(* Logix 5000 project; controller POA Emulate 5570 rev 30.12; software revision 30.00; part 4 of 6 *)
(* tags used below, declared in another part *)
   Chaskey_Message : DINT[256];
   Chaskey_mlen : DINT;
   Chaskey_MsgBitLen : DINT;
   Chaskey_round : DINT;
   Chaskey_tag : DINT[4];
   Date_time : DINT[7];
   OWF_Add_c : DINT;
   OWF_i : DINT;
   OWF_Input : DINT[17];
   OWF_InputLen : DINT;
   OWF_InputMaxInd : DINT;
   OWF_Result : DINT[17];
   POA_Chain_NM : DINT;
   POA_CKP : DINT[17];
   POA_i : DINT;
   POA_Ins_NM : DINT;
   POA_j : DINT;
   POA_k : DINT;
   POA_lr : DINT;
   POA_m : DINT;
   POA_Microsecond1 : DINT;
   POA_Microsecond2 : DINT;
   POA_MicrosecondABS : DINT;
   POA_OTS : SINT[256,256];
   POA_Pf : DINT[17];
   POA_Pf_Indx : DINT;
   POA_SC_Interval : DINT;
   POA_Second1 : DINT;
   POA_Second2 : DINT;
   POA_SecondABS : DINT;
   POA_SIG_i : DINT;
   POA_tag : DINT[4];
   POA_Vrf_Points : DINT[260,17];
   PRG_Counter : DINT[2];
   PRG_i : DINT;
   PRG_j : DINT;
   PRG_Res_Len : DINT;
   PRG_Result : DINT[128];
   SCAN_CYCLE_TIME : DINT;
   UOWHF_Add_c : DINT;
   UOWHF_Msg : DINT[17];
   UOWHF_Result : DINT[17];
   UOWHF_Vary_Message : DINT[3000];
   UOWHF_Vary_MsgLen : DINT;
   UOWHF_Ver : DINT;
(* MainProgram, continued *)

   		OWF_Add_c.1:=OWF_Result[1].31;
   		OWF_Result[1].31:=0;
   		OWF_Result[2]:=OWF_Result[2] + 102357735+OWF_Add_c;
   		OWF_Add_c.2:=OWF_Result[2].31;
   		OWF_Result[2].31:=0;
   		OWF_Result[3]:=OWF_Result[3] + 1548947751+OWF_Add_c;
   		OWF_Add_c.3:=OWF_Result[3].31;
   		OWF_Result[3].31:=0;
   		OWF_Result[4]:=OWF_Result[4] + 1541273950+OWF_Add_c;
   		OWF_Add_c.4:=OWF_Result[4].31;
   		OWF_Result[4].31:=0;
   		OWF_Result[5]:=OWF_Result[5] + 1965581916+OWF_Add_c;
   		OWF_Add_c.5:=OWF_Result[5].31;
   		OWF_Result[5].31:=0;
   		OWF_Result[6]:=OWF_Result[6] + 714783171+OWF_Add_c;
   		OWF_Add_c.6:=OWF_Result[6].31;
   		OWF_Result[6].31:=0;
   		OWF_Result[7]:=OWF_Result[7] + 952638591+OWF_Add_c;
   		OWF_Add_c.7:=OWF_Result[7].31;
   		OWF_Result[7].31:=0;
   		OWF_Result[8]:=OWF_Result[8] + 1892750752+OWF_Add_c;
   		OWF_Add_c.8:=OWF_Result[8].31;
   		OWF_Result[8].31:=0;
   	End_If;
   	If OWF_Input[7].[20] Then
   		OWF_Result[0]:=OWF_Result[0] + 1923601846+OWF_Add_c;
   		OWF_Add_c.0:=OWF_Result[0].31;
   		OWF_Result[0].31:=0;
   		OWF_Result[1]:=OWF_Result[1] + 431367542+OWF_Add_c;
   		OWF_Add_c.1:=OWF_Result[1].31;
   		OWF_Result[1].31:=0;
   		OWF_Result[2]:=OWF_Result[2] + 812772690+OWF_Add_c;
   		OWF_Add_c.2:=OWF_Result[2].31;
   		OWF_Result[2].31:=0;
   		OWF_Result[3]:=OWF_Result[3] + 1612004830+OWF_Add_c;
   		OWF_Add_c.3:=OWF_Result[3].31;
   		OWF_Result[3].31:=0;
   		OWF_Result[4]:=OWF_Result[4] + 1503607425+OWF_Add_c;
   		OWF_Add_c.4:=OWF_Result[4].31;
   		OWF_Result[4].31:=0;
   		OWF_Result[5]:=OWF_Result[5] + 257117095+OWF_Add_c;
   		OWF_Add_c.5:=OWF_Result[5].31;
   		OWF_Result[5].31:=0;
   		OWF_Result[6]:=OWF_Result[6] + 1165565758+OWF_Add_c;
   		OWF_Add_c.6:=OWF_Result[6].31;
   		OWF_Result[6].31:=0;
   		OWF_Result[7]:=OWF_Result[7] + 1791078952+OWF_Add_c;
   		OWF_Add_c.7:=OWF_Result[7].31;
   		OWF_Result[7].31:=0;
   		OWF_Result[8]:=OWF_Result[8] + 1316586480+OWF_Add_c;
   		OWF_Add_c.8:=OWF_Result[8].31;
   		OWF_Result[8].31:=0;
   	End_If;
   	If OWF_Input[7].[21] Then
   		OWF_Result[0]:=OWF_Result[0] + 1179130031+OWF_Add_c;
   		OWF_Add_c.0:=OWF_Result[0].31;
   		OWF_Result[0].31:=0;
   		OWF_Result[1]:=OWF_Result[1] + 1413483742+OWF_Add_c;
   		OWF_Add_c.1:=OWF_Result[1].31;
   		OWF_Result[1].31:=0;
   		OWF_Result[2]:=OWF_Result[2] + 2076538493+OWF_Add_c;
   		OWF_Add_c.2:=OWF_Result[2].31;
   		OWF_Result[2].31:=0;
   		OWF_Result[3]:=OWF_Result[3] + 415974763+OWF_Add_c;
   		OWF_Add_c.3:=OWF_Result[3].31;
   		OWF_Result[3].31:=0;
   		OWF_Result[4]:=OWF_Result[4] + 461079233+OWF_Add_c;
   		OWF_Add_c.4:=OWF_Result[4].31;
   		OWF_Result[4].31:=0;
   		OWF_Result[5]:=OWF_Result[5] + 207770264+OWF_Add_c;
   		OWF_Add_c.5:=OWF_Result[5].31;
   		OWF_Result[5].31:=0;
   		OWF_Result[6]:=OWF_Result[6] + 670532004+OWF_Add_c;
   		OWF_Add_c.6:=OWF_Result[6].31;
   		OWF_Result[6].31:=0;
   		OWF_Result[7]:=OWF_Result[7] + 164283060+OWF_Add_c;
   		OWF_Add_c.7:=OWF_Result[7].31;
   		OWF_Result[7].31:=0;
   		OWF_Result[8]:=OWF_Result[8] + 1512816438+OWF_Add_c;
   		OWF_Add_c.8:=OWF_Result[8].31;
   		OWF_Result[8].31:=0;
   	End_If;
   	If OWF_Input[7].[22] Then
   		OWF_Result[0]:=OWF_Result[0] + 1897360171+OWF_Add_c;
   		OWF_Add_c.0:=OWF_Result[0].31;
   		OWF_Result[0].31:=0;
   		OWF_Result[1]:=OWF_Result[1] + 1308779824+OWF_Add_c;
   		OWF_Add_c.1:=OWF_Result[1].31;
   		OWF_Result[1].31:=0;
   		OWF_Result[2]:=OWF_Result[2] + 1875593423+OWF_Add_c;
   		OWF_Add_c.2:=OWF_Result[2].31;
   		OWF_Result[2].31:=0;
   		OWF_Result[3]:=OWF_Result[3] + 571271217+OWF_Add_c;
   		OWF_Add_c.3:=OWF_Result[3].31;
   		OWF_Result[3].31:=0;
   		OWF_Result[4]:=OWF_Result[4] + 344940971+OWF_Add_c;
   		OWF_Add_c.4:=OWF_Result[4].31;
   		OWF_Result[4].31:=0;
   		OWF_Result[5]:=OWF_Result[5] + 75339231+OWF_Add_c;
   		OWF_Add_c.5:=OWF_Result[5].31;
   		OWF_Result[5].31:=0;
   		OWF_Result[6]:=OWF_Result[6] + 1428316860+OWF_Add_c;
   		OWF_Add_c.6:=OWF_Result[6].31;
   		OWF_Result[6].31:=0;
   		OWF_Result[7]:=OWF_Result[7] + 1811603075+OWF_Add_c;
   		OWF_Add_c.7:=OWF_Result[7].31;
   		OWF_Result[7].31:=0;
   		OWF_Result[8]:=OWF_Result[8] + 1679786029+OWF_Add_c;
   		OWF_Add_c.8:=OWF_Result[8].31;
   		OWF_Result[8].31:=0;
   	End_If;
   	If OWF_Input[7].[23] Then
   		OWF_Result[0]:=OWF_Result[0] + 271831917+OWF_Add_c;
   		OWF_Add_c.0:=OWF_Result[0].31;
   		OWF_Result[0].31:=0;
   		OWF_Result[1]:=OWF_Result[1] + 663117307+OWF_Add_c;
   		OWF_Add_c.1:=OWF_Result[1].31;
   		OWF_Result[1].31:=0;
   		OWF_Result[2]:=OWF_Result[2] + 1802435718+OWF_Add_c;
   		OWF_Add_c.2:=OWF_Result[2].31;
   		OWF_Result[2].31:=0;
   		OWF_Result[3]:=OWF_Result[3] + 585874673+OWF_Add_c;
   		OWF_Add_c.3:=OWF_Result[3].31;
   		OWF_Result[3].31:=0;
   		OWF_Result[4]:=OWF_Result[4] + 701698092+OWF_Add_c;
   		OWF_Add_c.4:=OWF_Result[4].31;
   		OWF_Result[4].31:=0;
   		OWF_Result[5]:=OWF_Result[5] + 1402770880+OWF_Add_c;
   		OWF_Add_c.5:=OWF_Result[5].31;
   		OWF_Result[5].31:=0;
   		OWF_Result[6]:=OWF_Result[6] + 452824658+OWF_Add_c;
   		OWF_Add_c.6:=OWF_Result[6].31;
   		OWF_Result[6].31:=0;
   		OWF_Result[7]:=OWF_Result[7] + 1400742763+OWF_Add_c;
   		OWF_Add_c.7:=OWF_Result[7].31;
   		OWF_Result[7].31:=0;
   		OWF_Result[8]:=OWF_Result[8] + 2073024045+OWF_Add_c;
   		OWF_Add_c.8:=OWF_Result[8].31;
   		OWF_Result[8].31:=0;
   	End_If;
   	If OWF_Input[7].[24] Then
   		OWF_Result[0]:=OWF_Result[0] + 1367845667+OWF_Add_c;
   		OWF_Add_c.0:=OWF_Result[0].31;
   		OWF_Result[0].31:=0;
   		OWF_Result[1]:=OWF_Result[1] + 1195094582+OWF_Add_c;
   		OWF_Add_c.1:=OWF_Result[1].31;
   		OWF_Result[1].31:=0;
   		OWF_Result[2]:=OWF_Result[2] + 494736933+OWF_Add_c;
   		OWF_Add_c.2:=OWF_Result[2].31;
   		OWF_Result[2].31:=0;
   		OWF_Result[3]:=OWF_Result[3] + 1875737261+OWF_Add_c;
   		OWF_Add_c.3:=OWF_Result[3].31;
   		OWF_Result[3].31:=0;
   		OWF_Result[4]:=OWF_Result[4] + 726339725+OWF_Add_c;
   		OWF_Add_c.4:=OWF_Result[4].31;
   		OWF_Result[4].31:=0;
   		OWF_Result[5]:=OWF_Result[5] + 1862851936+OWF_Add_c;
   		OWF_Add_c.5:=OWF_Result[5].31;
   		OWF_Result[5].31:=0;
   		OWF_Result[6]:=OWF_Result[6] + 296798862+OWF_Add_c;
   		OWF_Add_c.6:=OWF_Result[6].31;
   		OWF_Result[6].31:=0;
   		OWF_Result[7]:=OWF_Result[7] + 1485306441+OWF_Add_c;
   		OWF_Add_c.7:=OWF_Result[7].31;
   		OWF_Result[7].31:=0;
   		OWF_Result[8]:=OWF_Result[8] + 79244469+OWF_Add_c;
   		OWF_Add_c.8:=OWF_Result[8].31;
   		OWF_Result[8].31:=0;
   	End_If;
   	If OWF_Input[7].[25] Then
   		OWF_Result[0]:=OWF_Result[0] + 1748009068+OWF_Add_c;
   		OWF_Add_c.0:=OWF_Result[0].31;
   		OWF_Result[0].31:=0;
   		OWF_Result[1]:=OWF_Result[1] + 153673379+OWF_Add_c;
   		OWF_Add_c.1:=OWF_Result[1].31;
   		OWF_Result[1].31:=0;
   		OWF_Result[2]:=OWF_Result[2] + 1563899973+OWF_Add_c;
   		OWF_Add_c.2:=OWF_Result[2].31;
   		OWF_Result[2].31:=0;
   		OWF_Result[3]:=OWF_Result[3] + 210477071+OWF_Add_c;
   		OWF_Add_c.3:=OWF_Result[3].31;
   		OWF_Result[3].31:=0;
   		OWF_Result[4]:=OWF_Result[4] + 598591903+OWF_Add_c;
   		OWF_Add_c.4:=OWF_Result[4].31;
   		OWF_Result[4].31:=0;
   		OWF_Result[5]:=OWF_Result[5] + 889903791+OWF_Add_c;
   		OWF_Add_c.5:=OWF_Result[5].31;
   		OWF_Result[5].31:=0;
   		OWF_Result[6]:=OWF_Result[6] + 1087681228+OWF_Add_c;
   		OWF_Add_c.6:=OWF_Result[6].31;
   		OWF_Result[6].31:=0;
   		OWF_Result[7]:=OWF_Result[7] + 146945819+OWF_Add_c;
   		OWF_Add_c.7:=OWF_Result[7].31;
   		OWF_Result[7].31:=0;
   		OWF_Result[8]:=OWF_Result[8] + 658778953+OWF_Add_c;
   		OWF_Add_c.8:=OWF_Result[8].31;
   		OWF_Result[8].31:=0;
   	End_If;
   	If OWF_Input[7].[26] Then
   		OWF_Result[0]:=OWF_Result[0] + 1388889236+OWF_Add_c;
   		OWF_Add_c.0:=OWF_Result[0].31;
   		OWF_Result[0].31:=0;
   		OWF_Result[1]:=OWF_Result[1] + 1854230592+OWF_Add_c;
   		OWF_Add_c.1:=OWF_Result[1].31;
   		OWF_Result[1].31:=0;
   		OWF_Result[2]:=OWF_Result[2] + 1952659775+OWF_Add_c;
   		OWF_Add_c.2:=OWF_Result[2].31;
   		OWF_Result[2].31:=0;
   		OWF_Result[3]:=OWF_Result[3] + 693016622+OWF_Add_c;
   		OWF_Add_c.3:=OWF_Result[3].31;
   		OWF_Result[3].31:=0;
   		OWF_Result[4]:=OWF_Result[4] + 19961190+OWF_Add_c;
   		OWF_Add_c.4:=OWF_Result[4].31;
   		OWF_Result[4].31:=0;
   		OWF_Result[5]:=OWF_Result[5] + 1155238848+OWF_Add_c;
   		OWF_Add_c.5:=OWF_Result[5].31;
   		OWF_Result[5].31:=0;
   		OWF_Result[6]:=OWF_Result[6] + 1721973623+OWF_Add_c;
   		OWF_Add_c.6:=OWF_Result[6].31;
   		OWF_Result[6].31:=0;
   		OWF_Result[7]:=OWF_Result[7] + 1298626904+OWF_Add_c;
   		OWF_Add_c.7:=OWF_Result[7].31;
   		OWF_Result[7].31:=0;
   		OWF_Result[8]:=OWF_Result[8] + 704184103+OWF_Add_c;
   		OWF_Add_c.8:=OWF_Result[8].31;
   		OWF_Result[8].31:=0;
   	End_If;
   	If OWF_Input[7].[27] Then
   		OWF_Result[0]:=OWF_Result[0] + 1064559134+OWF_Add_c;
   		OWF_Add_c.0:=OWF_Result[0].31;
   		OWF_Result[0].31:=0;
   		OWF_Result[1]:=OWF_Result[1] + 628496468+OWF_Add_c;
   		OWF_Add_c.1:=OWF_Result[1].31;
   		OWF_Result[1].31:=0;
   		OWF_Result[2]:=OWF_Result[2] + 1741787667+OWF_Add_c;
   		OWF_Add_c.2:=OWF_Result[2].31;
   		OWF_Result[2].31:=0;
   		OWF_Result[3]:=OWF_Result[3] + 650880797+OWF_Add_c;
   		OWF_Add_c.3:=OWF_Result[3].31;
   		OWF_Result[3].31:=0;
   		OWF_Result[4]:=OWF_Result[4] + 927193641+OWF_Add_c;
   		OWF_Add_c.4:=OWF_Result[4].31;
   		OWF_Result[4].31:=0;
   		OWF_Result[5]:=OWF_Result[5] + 690779087+OWF_Add_c;
   		OWF_Add_c.5:=OWF_Result[5].31;
   		OWF_Result[5].31:=0;
   		OWF_Result[6]:=OWF_Result[6] + 1387171811+OWF_Add_c;
   		OWF_Add_c.6:=OWF_Result[6].31;
   		OWF_Result[6].31:=0;
   		OWF_Result[7]:=OWF_Result[7] + 1642242275+OWF_Add_c;
   		OWF_Add_c.7:=OWF_Result[7].31;
   		OWF_Result[7].31:=0;
   		OWF_Result[8]:=OWF_Result[8] + 750154437+OWF_Add_c;
   		OWF_Add_c.8:=OWF_Result[8].31;
   		OWF_Result[8].31:=0;
   	End_If;
   	If OWF_Input[7].[28] Then
   		OWF_Result[0]:=OWF_Result[0] + 1648370074+OWF_Add_c;
   		OWF_Add_c.0:=OWF_Result[0].31;
   		OWF_Result[0].31:=0;
   		OWF_Result[1]:=OWF_Result[1] + 242619355+OWF_Add_c;
   		OWF_Add_c.1:=OWF_Result[1].31;
   		OWF_Result[1].31:=0;
   		OWF_Result[2]:=OWF_Result[2] + 1874736599+OWF_Add_c;
   		OWF_Add_c.2:=OWF_Result[2].31;
   		OWF_Result[2].31:=0;
   		OWF_Result[3]:=OWF_Result[3] + 1413909693+OWF_Add_c;
   		OWF_Add_c.3:=OWF_Result[3].31;
   		OWF_Result[3].31:=0;
   		OWF_Result[4]:=OWF_Result[4] + 415302371+OWF_Add_c;
   		OWF_Add_c.4:=OWF_Result[4].31;
   		OWF_Result[4].31:=0;
   		OWF_Result[5]:=OWF_Result[5] + 2103173316+OWF_Add_c;
   		OWF_Add_c.5:=OWF_Result[5].31;
   		OWF_Result[5].31:=0;
   		OWF_Result[6]:=OWF_Result[6] + 317087375+OWF_Add_c;
   		OWF_Add_c.6:=OWF_Result[6].31;
   		OWF_Result[6].31:=0;
   		OWF_Result[7]:=OWF_Result[7] + 1550821217+OWF_Add_c;
   		OWF_Add_c.7:=OWF_Result[7].31;
   		OWF_Result[7].31:=0;
   		OWF_Result[8]:=OWF_Result[8] + 61155956+OWF_Add_c;
   		OWF_Add_c.8:=OWF_Result[8].31;
   		OWF_Result[8].31:=0;
   	End_If;
   	If OWF_Input[7].[29] Then
   		OWF_Result[0]:=OWF_Result[0] + 632604897+OWF_Add_c;
   		OWF_Add_c.0:=OWF_Result[0].31;
   		OWF_Result[0].31:=0;
   		OWF_Result[1]:=OWF_Result[1] + 1890179507+OWF_Add_c;
   		OWF_Add_c.1:=OWF_Result[1].31;
   		OWF_Result[1].31:=0;
   		OWF_Result[2]:=OWF_Result[2] + 1607995656+OWF_Add_c;
   		OWF_Add_c.2:=OWF_Result[2].31;
   		OWF_Result[2].31:=0;
   		OWF_Result[3]:=OWF_Result[3] + 1449206150+OWF_Add_c;
   		OWF_Add_c.3:=OWF_Result[3].31;
   		OWF_Result[3].31:=0;
   		OWF_Result[4]:=OWF_Result[4] + 402726737+OWF_Add_c;
   		OWF_Add_c.4:=OWF_Result[4].31;
   		OWF_Result[4].31:=0;
   		OWF_Result[5]:=OWF_Result[5] + 365091023+OWF_Add_c;
   		OWF_Add_c.5:=OWF_Result[5].31;
   		OWF_Result[5].31:=0;
   		OWF_Result[6]:=OWF_Result[6] + 1662601056+OWF_Add_c;
   		OWF_Add_c.6:=OWF_Result[6].31;
   		OWF_Result[6].31:=0;
   		OWF_Result[7]:=OWF_Result[7] + 1022070658+OWF_Add_c;
   		OWF_Add_c.7:=OWF_Result[7].31;
   		OWF_Result[7].31:=0;
   		OWF_Result[8]:=OWF_Result[8] + 49749052+OWF_Add_c;
   		OWF_Add_c.8:=OWF_Result[8].31;
   		OWF_Result[8].31:=0;
   	End_If;
   	If OWF_Input[7].[30] Then
   		OWF_Result[0]:=OWF_Result[0] + 1218340763+OWF_Add_c;
   		OWF_Add_c.0:=OWF_Result[0].31;
   		OWF_Result[0].31:=0;
   		OWF_Result[1]:=OWF_Result[1] + 1701757107+OWF_Add_c;
   		OWF_Add_c.1:=OWF_Result[1].31;
   		OWF_Result[1].31:=0;
   		OWF_Result[2]:=OWF_Result[2] + 1789117076+OWF_Add_c;
   		OWF_Add_c.2:=OWF_Result[2].31;
   		OWF_Result[2].31:=0;
   		OWF_Result[3]:=OWF_Result[3] + 963840108+OWF_Add_c;
   		OWF_Add_c.3:=OWF_Result[3].31;
   		OWF_Result[3].31:=0;
   		OWF_Result[4]:=OWF_Result[4] + 660620140+OWF_Add_c;
   		OWF_Add_c.4:=OWF_Result[4].31;
   		OWF_Result[4].31:=0;
   		OWF_Result[5]:=OWF_Result[5] + 983419398+OWF_Add_c;
   		OWF_Add_c.5:=OWF_Result[5].31;
   		OWF_Result[5].31:=0;
   		OWF_Result[6]:=OWF_Result[6] + 540791099+OWF_Add_c;
   		OWF_Add_c.6:=OWF_Result[6].31;
   		OWF_Result[6].31:=0;
   		OWF_Result[7]:=OWF_Result[7] + 2120149871+OWF_Add_c;
   		OWF_Add_c.7:=OWF_Result[7].31;
   		OWF_Result[7].31:=0;
   		OWF_Result[8]:=OWF_Result[8] + 1356988421+OWF_Add_c;
   		OWF_Add_c.8:=OWF_Result[8].31;
   		OWF_Result[8].31:=0;
   	End_If;
   	If OWF_Input[7].[31] Then
   		OWF_Result[0]:=OWF_Result[0] + 1135594880+OWF_Add_c;
   		OWF_Add_c.0:=OWF_Result[0].31;
   		OWF_Result[0].31:=0;
   		OWF_Result[1]:=OWF_Result[1] + 1430344149+OWF_Add_c;
   		OWF_Add_c.1:=OWF_Result[1].31;
   		OWF_Result[1].31:=0;
   		OWF_Result[2]:=OWF_Result[2] + 426577698+OWF_Add_c;
   		OWF_Add_c.2:=OWF_Result[2].31;
   		OWF_Result[2].31:=0;
   		OWF_Result[3]:=OWF_Result[3] + 34487438+OWF_Add_c;
   		OWF_Add_c.3:=OWF_Result[3].31;
   		OWF_Result[3].31:=0;
   		OWF_Result[4]:=OWF_Result[4] + 142555847+OWF_Add_c;
   		OWF_Add_c.4:=OWF_Result[4].31;
   		OWF_Result[4].31:=0;
   		OWF_Result[5]:=OWF_Result[5] + 380868128+OWF_Add_c;
   		OWF_Add_c.5:=OWF_Result[5].31;
   		OWF_Result[5].31:=0;
   		OWF_Result[6]:=OWF_Result[6] + 797337152+OWF_Add_c;
   		OWF_Add_c.6:=OWF_Result[6].31;
   		OWF_Result[6].31:=0;
   		OWF_Result[7]:=OWF_Result[7] + 1153550956+OWF_Add_c;
   		OWF_Add_c.7:=OWF_Result[7].31;
   		OWF_Result[7].31:=0;
   		OWF_Result[8]:=OWF_Result[8] + 2080693926+OWF_Add_c;
   		OWF_Add_c.8:=OWF_Result[8].31;
   		OWF_Result[8].31:=0;
   	End_If;
   
   	OWF_Result[OWF_InputMaxInd]:=OWF_Result[OWF_InputMaxInd] and 16#FF; //clear high bit
   
END_ROUTINE

ROUTINE Improved_OWF   (* structured text *)
   
   
   JSR(OWF_Init);
   JSR(If256);
END_ROUTINE

ROUTINE MainRoutine   (* ladder *)
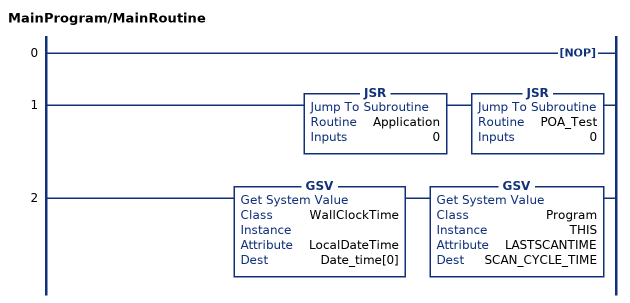
   0: NOP();
   1: JSR(Application,0)JSR(POA_Test,0);
   2: GSV(WallClockTime,,LocalDateTime,Date_time[0])GSV(Program,THIS,LASTSCANTIME,SCAN_CYCLE_TIME);
END_ROUTINE

ROUTINE OWF_Init   (* structured text *)
   OWF_InputLen:=255;  //bits of input.
   OWF_InputMaxInd:=8;  //maximum index for dints which store the bits of input.
   
   
   For OWF_i:=0 to OWF_InputMaxInd by 1 do
   	OWF_Result[OWF_i]:=0;
   End_For;
   
   
END_ROUTINE

ROUTINE POA_PF_Init   (* structured text *)
   	POA_lr :=8;  //256 bits
   
   	POA_SC_Interval:=8388608;  // 2^23;
   
   	POA_Pf_Indx:= 64;  //the number of passwords in a OWF chain
   
   
END_ROUTINE

ROUTINE POA_ProofGeneration   (* structured text *)
   
   	JSR(POA_PF_Init);
   
   	POA_Second2:=Date_time[5];  //second
   	POA_Microsecond2:=Date_time[6];  //Microsecond
   
   	POA_SecondABS:=ABS(POA_Second2 - POA_Second1);
   	POA_MicrosecondABS:=ABS(POA_Microsecond2-POA_Microsecond1);
   	if (POA_SecondABS*1000000+POA_MicrosecondABS)>60000000 then
   		//There was an attack, rasise an alarm....60000000 is 60 seconds
   	end_if;
   
   	//run chaskey to verify the MAC
   	Chaskey_Message[0]:= POA_Pf_Indx;
   	Chaskey_Message[1] := POA_Chain_NM;
   	Chaskey_Message[2] := POA_Ins_NM;
   	Chaskey_Message[3]:=POA_Second1;   //Add time to message to compute MAC.
   	Chaskey_Message[4]:=POA_Microsecond1;   //Add time to message to compute MAC.
   	//Chaskey_m_len:=1696;
   	Chaskey_round:=7;
   	Chaskey_mlen:=4;
   	Chaskey_MsgBitLen:=160;
   	JSR(CHASKEY_128);
   
   	If POA_tag[3]<>Chaskey_tag[3] OR POA_tag[2]<> Chaskey_tag[2]  OR POA_tag[1]<> Chaskey_tag[1] OR POA_tag[0]<> Chaskey_tag[0] then
   		//There was an attack, rasise an alarm....
   	end_if;
   
   	//use PRG to generate the head node
   	PRG_Counter[0]:= POA_Ins_NM;
   	PRG_Counter[1]:= POA_Chain_NM + POA_lr;
   	JSR(PRG_PRF_CHASKEY);
   	//256-bits result of MAC assign to checkpoint
   	for POA_i:=0 to 7 by 1 do
   		POA_CKP[POA_i]:=PRG_Result[POA_i];
   	end_for;
   	//use OWF to generate every check point
   	OWF_Input[0]:=POA_CKP[0];
   	OWF_Input[1]:=POA_CKP[1];
   	OWF_Input[2]:=POA_CKP[2];
   	OWF_Input[3]:=POA_CKP[3];
   	OWF_Input[4]:=POA_CKP[4];
   	OWF_Input[5]:=POA_CKP[5];
   	OWF_Input[6]:=POA_CKP[6];
   	OWF_Input[7]:=POA_CKP[7];
   	OWF_Input[8]:=POA_CKP[8];
   
   	for POA_j:=0 to POA_Pf_Indx by 1 do
   		JSR(Improved_OWF);
   			OWF_Input[0]:=OWF_Result[0];
   			OWF_Input[1]:=OWF_Result[1];
   			OWF_Input[2]:=OWF_Result[2];
   			OWF_Input[3]:=OWF_Result[3];
   			OWF_Input[4]:=OWF_Result[4];
   			OWF_Input[5]:=OWF_Result[5];
   			OWF_Input[6]:=OWF_Result[6];
   			OWF_Input[7]:=OWF_Result[7];
   			OWF_Input[8]:=OWF_Result[8];
   	end_for;
   
   	for POA_j:=0 to 7 by 1 do
   		POA_Pf[POA_j]:= OWF_Result[POA_j];
   	end_for;
   
   	POA_Pf_Indx:=POA_Pf_Indx -1;
   
   	if (POA_Pf_Indx=1) and (POA_Chain_NM=2139095040) then
   
   		JSR(POA_Replenishment);
   	end_if;
   
   	//update check point's index..
   	if POA_Pf_Indx-1 = 1 then
   		if POA_Chain_NM<>256 then	// the chain is not used out
   			POA_Chain_NM:=POA_Chain_NM+POA_SC_Interval;
   		end_if;
   	end_if;
   
   	POA_Second1:=Date_time[5];
   	POA_Microsecond1:=Date_time[6];
   
   	Chaskey_Message[0]:= POA_Pf_Indx;
   	Chaskey_Message[1] := POA_Chain_NM;
   	Chaskey_Message[2] := POA_Ins_NM;
   	Chaskey_Message[3]:=POA_Second1;   //Add time to message to compute MAC.
   	Chaskey_Message[4]:=POA_Microsecond1;   //Add time to message to compute MAC.
   	Chaskey_MsgBitLen:=160;  //5*32 bits.
   	Chaskey_mlen:=4;
   	Chaskey_round:=7;
   	JSR(CHASKEY_128);
   
   	POA_tag[3]:=Chaskey_tag[3] ;
   	POA_tag[2]:=Chaskey_tag[2]  ;
   	POA_tag[1]:=Chaskey_tag[1] ;
   	POA_tag[0]:=Chaskey_tag[0] ;
   
   	//POA_time1:=GSV(WallClockTime,LocalDateTime,Date_time[6]);
   
   	// clear the credentials
   	for POA_j:=0 to 7 by 1 do
   		POA_CKP[POA_j]:=0;
   		PRG_Result[POA_j]:=0;
   	end_for;
   
   
   
END_ROUTINE

ROUTINE POA_ReInit   (* structured text *)
   //POA_PRG_Indx for replenishment
   
   
   	POA_Ins_NM:= POA_Ins_NM+1;  //compute a new instance.
   
   	POA_Chain_NM :=0;   //the number of OWF sub-chain
   
   
   
   	UOWHF_Ver:=0;
   
   
   	JSR(POA_PF_Init);
   
   
   
   
   
END_ROUTINE

ROUTINE POA_Replenishment   (* structured text *)
   
   JSR(POA_ReInit);
   
   
   //compute all the tail of each OWF chain.
   
   for POA_m:=0 to 255 by 1 do
   //POA_k:=0 to POA_SC_Interval*255 by POA_SC_Interval do
   	//use PRG to generate the head node
   	PRG_Counter[0]:= POA_Ins_NM;
   	PRG_Counter[1]:= POA_Chain_NM + POA_lr;
   
   	JSR(PRG_PRF_CHASKEY);
   
   	for POA_i:=0 to 8 by 1 do   //256-bits result of MAC assign to checkpoint.
   
   		//POA_CKP[POA_i]:=PRG_Result[POA_i];
   		POA_CKP[POA_i]:=65535;
   
   	end_for;
   
   	OWF_Input[0]:=POA_CKP[0];
   	OWF_Input[1]:=POA_CKP[1];
   	OWF_Input[2]:=POA_CKP[2];
   	OWF_Input[3]:=POA_CKP[3];
   	OWF_Input[4]:=POA_CKP[4];
   	OWF_Input[5]:=POA_CKP[5];
   	OWF_Input[6]:=POA_CKP[6];
   	OWF_Input[7]:=POA_CKP[7];
   	OWF_Input[8]:=POA_CKP[8];
   
   	for POA_j:=0 to POA_Pf_Indx by 1 do   //compute the tail of one OWF chain.
   		JSR(Improved_OWF);
   		OWF_Input[0]:=OWF_Result[0];
   		OWF_Input[1]:=OWF_Result[1];
   		OWF_Input[2]:=OWF_Result[2];
   		OWF_Input[3]:=OWF_Result[3];
   		OWF_Input[4]:=OWF_Result[4];
   		OWF_Input[5]:=OWF_Result[5];
   		OWF_Input[6]:=OWF_Result[6];
   		OWF_Input[7]:=OWF_Result[7];
   		OWF_Input[8]:=POA_CKP[8];
   	end_for;
   
   	for POA_j:=0 to 8 by 1 do  //store all the tail.
   		POA_Vrf_Points[POA_m,POA_j]:= OWF_Result[POA_j];
   	end_for;
   	POA_Chain_NM:=POA_Chain_NM+POA_SC_Interval;
   
   end_for;
   
   
   //all tail as input message, compute the hash of all tail.
   UOWHF_Vary_MsgLen:=2047;  //256*8 Dints
   for POA_j:=0 to 255 by 1 do   //assign the tail value to Hash_Msg[].
   	for POA_i:=0 to 8 by 1 do
   		UOWHF_Vary_Message[POA_i+8*POA_j]:=POA_Vrf_Points[POA_j,POA_i];
   	end_for;
   end_for;
   JSR(UOWHF_Vary);  //gain the Hash result with 128 bits.
   
   
   
   
   // compute OTS using the heads of the last protocol instance...................
   POA_k:=0;
   POA_SIG_i:=0;
   for POA_i:=0 to 3 by 1 do
   	for POA_j:=0 to 31 by 1 do
   		if OWF_Result[POA_i].[POA_j] then  //if bit is 1, choose the second head as sk.
   			PRG_Counter[0]:= POA_Ins_NM-1;
   			PRG_Counter[1]:= 2*POA_k+POA_SC_Interval + POA_lr;
   
   			JSR(PRG_PRF_CHASKEY);
   
   
   		else
   			PRG_Counter[0]:= POA_Ins_NM-1;
   			PRG_Counter[1]:= 2*POA_k + POA_lr;
   
   			JSR(PRG_PRF_CHASKEY);
   		end_if;
   
   		for POA_m:=0 to 7 by 1 do
   			POA_OTS[POA_SIG_i,POA_m]:=PRG_Result[POA_m]; //store all the result of OTS.
   		end_for;
   	POA_k:=POA_k+POA_SC_Interval;
   	POA_SIG_i:=POA_SIG_i+1;
   	end_for;
   end_for;
   
   
   // clear the credentials
   for POA_j:=0 to 8 by 1 do
   	POA_CKP[POA_j]:=0;
   	PRG_Result[POA_j]:=0;
   end_for;
   
   
   
END_ROUTINE

ROUTINE POA_Test   (* structured text *)
   If S:FS Then
   	jsr(POA_PF_Init);
   
   
   End_If;
   
   //JSR(POA_ProofGeneration);
   JSR(POA_Replenishment);
END_ROUTINE

ROUTINE PRG_PRF_CHASKEY   (* structured text *)
   // init PRG_Count[0] and PRG_Count[1] during application.. for PRF.. they could be any values
   //For PRG application, PRG_Count[0] defines the output length (i.e., the number of 64-bit, e.g., 128-bit output, PRG_Count[0]:=2)
   
   
   JSR(PRG_PRF_Init);
   PRG_j:=0;
   For PRG_i:=0 to PRG_Res_Len by 1 do
   	Chaskey_Message[0]:=PRG_Counter[0]; //Upper bits of current plaintext
   	Chaskey_Message[1]:=PRG_Counter[1];  //Lower bits of current plaintext
   	Chaskey_Message[2]:=PRG_Counter[0]; //Upper bits of current plaintext
   	Chaskey_Message[3]:=PRG_Counter[1];  //Lower bits of current plaintext
   	JSR(CHASKEY_128);
   	PRG_Result[PRG_j]:=Chaskey_tag[0];
   	PRG_Result[PRG_j+1]:=Chaskey_tag[1];
   	PRG_Result[PRG_j+2]:=Chaskey_tag[2];
   	PRG_Result[PRG_j+3]:=Chaskey_tag[3];
   
   	PRG_j:=PRG_j+4;
   
   End_For;
   
   JSR(CHASKEY_ClearKey);
   
END_ROUTINE

ROUTINE PRG_PRF_Init   (* structured text *)
   //initialize version
   
   
   Chaskey_round:=11;
   PRG_j:=0;
   PRG_Res_Len :=  (PRG_Counter[0] AND 16#0000ffff)-1;
   
   JSR(CHASKEY_Init);
END_ROUTINE

ROUTINE UOWHF   (* structured text *)
   
   
   
   
    JSR(UOWHF_Init);
   
   
   
   
   		Case UOWHF_Ver OF
   		0:
   			JSR(UOWHF_If256);
   		1:
   
   		2:
   
   		End_Case;
   
   
END_ROUTINE

ROUTINE UOWHF_If256   (* structured text *)
   	If UOWHF_Msg[0].[0] Then
   		UOWHF_Result[0]:=UOWHF_Result[0] + 572632243+UOWHF_Add_c;
   		UOWHF_Add_c.0:=UOWHF_Result[0].31;
   		UOWHF_Result[0].31:=0;
   		UOWHF_Result[1]:=UOWHF_Result[1] + 477137765+UOWHF_Add_c;
   		UOWHF_Add_c.1:=UOWHF_Result[1].31;
   		UOWHF_Result[1].31:=0;
   		UOWHF_Result[2]:=UOWHF_Result[2] + 550157017+UOWHF_Add_c;
   		UOWHF_Add_c.2:=UOWHF_Result[2].31;
   		UOWHF_Result[2].31:=0;
   		UOWHF_Result[3]:=UOWHF_Result[3] + 245297039+UOWHF_Add_c;
   		UOWHF_Add_c.3:=UOWHF_Result[3].31;
   		UOWHF_Result[3].31:=0;
   		UOWHF_Result[4]:=UOWHF_Result[4] + 890022153+UOWHF_Add_c;
   		UOWHF_Add_c.4:=UOWHF_Result[4].31;
   		UOWHF_Result[4].31:=0;
   	End_If;
   	If UOWHF_Msg[0].[1] Then
   		UOWHF_Result[0]:=UOWHF_Result[0] + 1377061044+UOWHF_Add_c;
   		UOWHF_Add_c.0:=UOWHF_Result[0].31;
   		UOWHF_Result[0].31:=0;
   		UOWHF_Result[1]:=UOWHF_Result[1] + 1295766427+UOWHF_Add_c;
   		UOWHF_Add_c.1:=UOWHF_Result[1].31;
   		UOWHF_Result[1].31:=0;
   		UOWHF_Result[2]:=UOWHF_Result[2] + 1302731282+UOWHF_Add_c;
   		UOWHF_Add_c.2:=UOWHF_Result[2].31;
   		UOWHF_Result[2].31:=0;
   		UOWHF_Result[3]:=UOWHF_Result[3] + 560246492+UOWHF_Add_c;
   		UOWHF_Add_c.3:=UOWHF_Result[3].31;
   		UOWHF_Result[3].31:=0;
   		UOWHF_Result[4]:=UOWHF_Result[4] + 148872358+UOWHF_Add_c;
   		UOWHF_Add_c.4:=UOWHF_Result[4].31;
   		UOWHF_Result[4].31:=0;
   	End_If;
   	If UOWHF_Msg[0].[2] Then
   		UOWHF_Result[0]:=UOWHF_Result[0] + 1840006150+UOWHF_Add_c;
   		UOWHF_Add_c.0:=UOWHF_Result[0].31;
   		UOWHF_Result[0].31:=0;
   		UOWHF_Result[1]:=UOWHF_Result[1] + 445834309+UOWHF_Add_c;
   		UOWHF_Add_c.1:=UOWHF_Result[1].31;
   		UOWHF_Result[1].31:=0;
   		UOWHF_Result[2]:=UOWHF_Result[2] + 927236896+UOWHF_Add_c;
   		UOWHF_Add_c.2:=UOWHF_Result[2].31;
   		UOWHF_Result[2].31:=0;
   		UOWHF_Result[3]:=UOWHF_Result[3] + 47182984+UOWHF_Add_c;
   		UOWHF_Add_c.3:=UOWHF_Result[3].31;
   		UOWHF_Result[3].31:=0;
   		UOWHF_Result[4]:=UOWHF_Result[4] + 50959418+UOWHF_Add_c;
   		UOWHF_Add_c.4:=UOWHF_Result[4].31;
   		UOWHF_Result[4].31:=0;
   	End_If;
   	If UOWHF_Msg[0].[3] Then
   		UOWHF_Result[0]:=UOWHF_Result[0] + 308042492+UOWHF_Add_c;
   		UOWHF_Add_c.0:=UOWHF_Result[0].31;
   		UOWHF_Result[0].31:=0;
   		UOWHF_Result[1]:=UOWHF_Result[1] + 822181770+UOWHF_Add_c;
   		UOWHF_Add_c.1:=UOWHF_Result[1].31;
   		UOWHF_Result[1].31:=0;
   		UOWHF_Result[2]:=UOWHF_Result[2] + 847762969+UOWHF_Add_c;
   		UOWHF_Add_c.2:=UOWHF_Result[2].31;
   		UOWHF_Result[2].31:=0;
   		UOWHF_Result[3]:=UOWHF_Result[3] + 1102323899+UOWHF_Add_c;
   		UOWHF_Add_c.3:=UOWHF_Result[3].31;
   		UOWHF_Result[3].31:=0;
   		UOWHF_Result[4]:=UOWHF_Result[4] + 606857113+UOWHF_Add_c;
   		UOWHF_Add_c.4:=UOWHF_Result[4].31;
   		UOWHF_Result[4].31:=0;
   	End_If;
   	If UOWHF_Msg[0].[4] Then
   		UOWHF_Result[0]:=UOWHF_Result[0] + 1879838005+UOWHF_Add_c;
   		UOWHF_Add_c.0:=UOWHF_Result[0].31;
   		UOWHF_Result[0].31:=0;
   		UOWHF_Result[1]:=UOWHF_Result[1] + 289434158+UOWHF_Add_c;
   		UOWHF_Add_c.1:=UOWHF_Result[1].31;
   		UOWHF_Result[1].31:=0;
   		UOWHF_Result[2]:=UOWHF_Result[2] + 2129379257+UOWHF_Add_c;
   		UOWHF_Add_c.2:=UOWHF_Result[2].31;
   		UOWHF_Result[2].31:=0;
   		UOWHF_Result[3]:=UOWHF_Result[3] + 1362062997+UOWHF_Add_c;
   		UOWHF_Add_c.3:=UOWHF_Result[3].31;
   		UOWHF_Result[3].31:=0;
   		UOWHF_Result[4]:=UOWHF_Result[4] + 1863755322+UOWHF_Add_c;
   		UOWHF_Add_c.4:=UOWHF_Result[4].31;
   		UOWHF_Result[4].31:=0;
   	End_If;
   	If UOWHF_Msg[0].[5] Then
   		UOWHF_Result[0]:=UOWHF_Result[0] + 1955367670+UOWHF_Add_c;
   		UOWHF_Add_c.0:=UOWHF_Result[0].31;
   		UOWHF_Result[0].31:=0;
   		UOWHF_Result[1]:=UOWHF_Result[1] + 126312607+UOWHF_Add_c;
   		UOWHF_Add_c.1:=UOWHF_Result[1].31;
   		UOWHF_Result[1].31:=0;
   		UOWHF_Result[2]:=UOWHF_Result[2] + 1694646926+UOWHF_Add_c;
   		UOWHF_Add_c.2:=UOWHF_Result[2].31;
   		UOWHF_Result[2].31:=0;
   		UOWHF_Result[3]:=UOWHF_Result[3] + 1429674455+UOWHF_Add_c;
   		UOWHF_Add_c.3:=UOWHF_Result[3].31;
   		UOWHF_Result[3].31:=0;
   		UOWHF_Result[4]:=UOWHF_Result[4] + 1469336309+UOWHF_Add_c;
   		UOWHF_Add_c.4:=UOWHF_Result[4].31;
   		UOWHF_Result[4].31:=0;
   	End_If;
   	If UOWHF_Msg[0].[6] Then
   		UOWHF_Result[0]:=UOWHF_Result[0] + 1633958070+UOWHF_Add_c;
   		UOWHF_Add_c.0:=UOWHF_Result[0].31;
   		UOWHF_Result[0].31:=0;
   		UOWHF_Result[1]:=UOWHF_Result[1] + 538621445+UOWHF_Add_c;
   		UOWHF_Add_c.1:=UOWHF_Result[1].31;
   		UOWHF_Result[1].31:=0;
   		UOWHF_Result[2]:=UOWHF_Result[2] + 2019575413+UOWHF_Add_c;
   		UOWHF_Add_c.2:=UOWHF_Result[2].31;
   		UOWHF_Result[2].31:=0;
   		UOWHF_Result[3]:=UOWHF_Result[3] + 995352028+UOWHF_Add_c;
   		UOWHF_Add_c.3:=UOWHF_Result[3].31;
   		UOWHF_Result[3].31:=0;
   		UOWHF_Result[4]:=UOWHF_Result[4] + 381457758+UOWHF_Add_c;
   		UOWHF_Add_c.4:=UOWHF_Result[4].31;
   		UOWHF_Result[4].31:=0;
   	End_If;
   	If UOWHF_Msg[0].[7] Then
   		UOWHF_Result[0]:=UOWHF_Result[0] + 357837682+UOWHF_Add_c;
   		UOWHF_Add_c.0:=UOWHF_Result[0].31;
   		UOWHF_Result[0].31:=0;
   		UOWHF_Result[1]:=UOWHF_Result[1] + 1524722817+UOWHF_Add_c;
   		UOWHF_Add_c.1:=UOWHF_Result[1].31;
   		UOWHF_Result[1].31:=0;
   		UOWHF_Result[2]:=UOWHF_Result[2] + 504152330+UOWHF_Add_c;
   		UOWHF_Add_c.2:=UOWHF_Result[2].31;
   		UOWHF_Result[2].31:=0;
   		UOWHF_Result[3]:=UOWHF_Result[3] + 1761625815+UOWHF_Add_c;
   		UOWHF_Add_c.3:=UOWHF_Result[3].31;
   		UOWHF_Result[3].31:=0;
   		UOWHF_Result[4]:=UOWHF_Result[4] + 944307141+UOWHF_Add_c;
   		UOWHF_Add_c.4:=UOWHF_Result[4].31;
   		UOWHF_Result[4].31:=0;
   	End_If;
   	If UOWHF_Msg[0].[8] Then
   		UOWHF_Result[0]:=UOWHF_Result[0] + 367007339+UOWHF_Add_c;
   		UOWHF_Add_c.0:=UOWHF_Result[0].31;
   		UOWHF_Result[0].31:=0;
   		UOWHF_Result[1]:=UOWHF_Result[1] + 1692729942+UOWHF_Add_c;
   		UOWHF_Add_c.1:=UOWHF_Result[1].31;
   		UOWHF_Result[1].31:=0;
   		UOWHF_Result[2]:=UOWHF_Result[2] + 2007351861+UOWHF_Add_c;
   		UOWHF_Add_c.2:=UOWHF_Result[2].31;
   		UOWHF_Result[2].31:=0;
   		UOWHF_Result[3]:=UOWHF_Result[3] + 1998537115+UOWHF_Add_c;
   		UOWHF_Add_c.3:=UOWHF_Result[3].31;
   		UOWHF_Result[3].31:=0;
   		UOWHF_Result[4]:=UOWHF_Result[4] + 538473612+UOWHF_Add_c;
   		UOWHF_Add_c.4:=UOWHF_Result[4].31;
   		UOWHF_Result[4].31:=0;
   	End_If;
   	If UOWHF_Msg[0].[9] Then
   		UOWHF_Result[0]:=UOWHF_Result[0] + 693038975+UOWHF_Add_c;
   		UOWHF_Add_c.0:=UOWHF_Result[0].31;
   		UOWHF_Result[0].31:=0;
   		UOWHF_Result[1]:=UOWHF_Result[1] + 1580596029+UOWHF_Add_c;
   		UOWHF_Add_c.1:=UOWHF_Result[1].31;
   		UOWHF_Result[1].31:=0;
   		UOWHF_Result[2]:=UOWHF_Result[2] + 2114924986+UOWHF_Add_c;
   		UOWHF_Add_c.2:=UOWHF_Result[2].31;
   		UOWHF_Result[2].31:=0;
   		UOWHF_Result[3]:=UOWHF_Result[3] + 1534063000+UOWHF_Add_c;
   		UOWHF_Add_c.3:=UOWHF_Result[3].31;
   		UOWHF_Result[3].31:=0;
   		UOWHF_Result[4]:=UOWHF_Result[4] + 1027147997+UOWHF_Add_c;
   		UOWHF_Add_c.4:=UOWHF_Result[4].31;
   		UOWHF_Result[4].31:=0;
   	End_If;
   	If UOWHF_Msg[0].[10] Then
   		UOWHF_Result[0]:=UOWHF_Result[0] + 817852360+UOWHF_Add_c;
   		UOWHF_Add_c.0:=UOWHF_Result[0].31;
   		UOWHF_Result[0].31:=0;
   		UOWHF_Result[1]:=UOWHF_Result[1] + 1240911531+UOWHF_Add_c;
   		UOWHF_Add_c.1:=UOWHF_Result[1].31;
   		UOWHF_Result[1].31:=0;
   		UOWHF_Result[2]:=UOWHF_Result[2] + 326514746+UOWHF_Add_c;
   		UOWHF_Add_c.2:=UOWHF_Result[2].31;
   		UOWHF_Result[2].31:=0;
   		UOWHF_Result[3]:=UOWHF_Result[3] + 1232608017+UOWHF_Add_c;
   		UOWHF_Add_c.3:=UOWHF_Result[3].31;
   		UOWHF_Result[3].31:=0;
   		UOWHF_Result[4]:=UOWHF_Result[4] + 28043263+UOWHF_Add_c;
   		UOWHF_Add_c.4:=UOWHF_Result[4].31;
   		UOWHF_Result[4].31:=0;
   	End_If;
   	If UOWHF_Msg[0].[11] Then
   		UOWHF_Result[0]:=UOWHF_Result[0] + 1640483064+UOWHF_Add_c;
   		UOWHF_Add_c.0:=UOWHF_Result[0].31;
   		UOWHF_Result[0].31:=0;
   		UOWHF_Result[1]:=UOWHF_Result[1] + 10392502+UOWHF_Add_c;
   		UOWHF_Add_c.1:=UOWHF_Result[1].31;
   		UOWHF_Result[1].31:=0;
   		UOWHF_Result[2]:=UOWHF_Result[2] + 1284374523+UOWHF_Add_c;
   		UOWHF_Add_c.2:=UOWHF_Result[2].31;
   		UOWHF_Result[2].31:=0;
   		UOWHF_Result[3]:=UOWHF_Result[3] + 1057415504+UOWHF_Add_c;
   		UOWHF_Add_c.3:=UOWHF_Result[3].31;
   		UOWHF_Result[3].31:=0;
   		UOWHF_Result[4]:=UOWHF_Result[4] + 79887159+UOWHF_Add_c;
   		UOWHF_Add_c.4:=UOWHF_Result[4].31;
   		UOWHF_Result[4].31:=0;
   	End_If;
   	If UOWHF_Msg[0].[12] Then
   		UOWHF_Result[0]:=UOWHF_Result[0] + 372752318+UOWHF_Add_c;
   		UOWHF_Add_c.0:=UOWHF_Result[0].31;
   		UOWHF_Result[0].31:=0;
   		UOWHF_Result[1]:=UOWHF_Result[1] + 858061594+UOWHF_Add_c;
   		UOWHF_Add_c.1:=UOWHF_Result[1].31;
   		UOWHF_Result[1].31:=0;
   		UOWHF_Result[2]:=UOWHF_Result[2] + 1568496385+UOWHF_Add_c;
   		UOWHF_Add_c.2:=UOWHF_Result[2].31;
   		UOWHF_Result[2].31:=0;
   		UOWHF_Result[3]:=UOWHF_Result[3] + 1501186385+UOWHF_Add_c;